(* Logix 5000 project; controller POA Emulate 5570 rev 30.12; software revision 30.00; part 6 of 6 *)
(* tags used below, declared in another part *)
   UOWHF_Add_c : DINT;
   UOWHF_i : DINT;
   UOWHF_InputLen : DINT;
   UOWHF_InputMaxInd : DINT;
   UOWHF_Msg : DINT[17];
   UOWHF_OutputMaxInd : DINT;
   UOWHF_Result : DINT[17];
   UOWHF_Vary_BlkNum : DINT;
   UOWHF_Vary_i : DINT;
   UOWHF_Vary_j : DINT;
   UOWHF_Vary_Message : DINT[3000];
   UOWHF_Vary_MsgLen : DINT;
   UOWHF_Vary_z : DINT;
   UOWHF_VaryLen : DINT;
   UOWHF_Ver : DINT;
(* MainProgram, continued *)

   		UOWHF_Result[0].31:=0;
   		UOWHF_Result[1]:=UOWHF_Result[1] + 1000119182+UOWHF_Add_c;
   		UOWHF_Add_c.1:=UOWHF_Result[1].31;
   		UOWHF_Result[1].31:=0;
   		UOWHF_Result[2]:=UOWHF_Result[2] + 1408193498+UOWHF_Add_c;
   		UOWHF_Add_c.2:=UOWHF_Result[2].31;
   		UOWHF_Result[2].31:=0;
   		UOWHF_Result[3]:=UOWHF_Result[3] + 758141530+UOWHF_Add_c;
   		UOWHF_Add_c.3:=UOWHF_Result[3].31;
   		UOWHF_Result[3].31:=0;
   		UOWHF_Result[4]:=UOWHF_Result[4] + 113758068+UOWHF_Add_c;
   		UOWHF_Add_c.4:=UOWHF_Result[4].31;
   		UOWHF_Result[4].31:=0;
   	End_If;
   	If UOWHF_Msg[7].[27] Then
   		UOWHF_Result[0]:=UOWHF_Result[0] + 86421407+UOWHF_Add_c;
   		UOWHF_Add_c.0:=UOWHF_Result[0].31;
   		UOWHF_Result[0].31:=0;
   		UOWHF_Result[1]:=UOWHF_Result[1] + 209732804+UOWHF_Add_c;
   		UOWHF_Add_c.1:=UOWHF_Result[1].31;
   		UOWHF_Result[1].31:=0;
   		UOWHF_Result[2]:=UOWHF_Result[2] + 502288861+UOWHF_Add_c;
   		UOWHF_Add_c.2:=UOWHF_Result[2].31;
   		UOWHF_Result[2].31:=0;
   		UOWHF_Result[3]:=UOWHF_Result[3] + 1399545115+UOWHF_Add_c;
   		UOWHF_Add_c.3:=UOWHF_Result[3].31;
   		UOWHF_Result[3].31:=0;
   		UOWHF_Result[4]:=UOWHF_Result[4] + 871725095+UOWHF_Add_c;
   		UOWHF_Add_c.4:=UOWHF_Result[4].31;
   		UOWHF_Result[4].31:=0;
   	End_If;
   	If UOWHF_Msg[7].[28] Then
   		UOWHF_Result[0]:=UOWHF_Result[0] + 2145748906+UOWHF_Add_c;
   		UOWHF_Add_c.0:=UOWHF_Result[0].31;
   		UOWHF_Result[0].31:=0;
   		UOWHF_Result[1]:=UOWHF_Result[1] + 750367767+UOWHF_Add_c;
   		UOWHF_Add_c.1:=UOWHF_Result[1].31;
   		UOWHF_Result[1].31:=0;
   		UOWHF_Result[2]:=UOWHF_Result[2] + 52958798+UOWHF_Add_c;
   		UOWHF_Add_c.2:=UOWHF_Result[2].31;
   		UOWHF_Result[2].31:=0;
   		UOWHF_Result[3]:=UOWHF_Result[3] + 299422686+UOWHF_Add_c;
   		UOWHF_Add_c.3:=UOWHF_Result[3].31;
   		UOWHF_Result[3].31:=0;
   		UOWHF_Result[4]:=UOWHF_Result[4] + 308572882+UOWHF_Add_c;
   		UOWHF_Add_c.4:=UOWHF_Result[4].31;
   		UOWHF_Result[4].31:=0;
   	End_If;
   	If UOWHF_Msg[7].[29] Then
   		UOWHF_Result[0]:=UOWHF_Result[0] + 470166861+UOWHF_Add_c;
   		UOWHF_Add_c.0:=UOWHF_Result[0].31;
   		UOWHF_Result[0].31:=0;
   		UOWHF_Result[1]:=UOWHF_Result[1] + 415982775+UOWHF_Add_c;
   		UOWHF_Add_c.1:=UOWHF_Result[1].31;
   		UOWHF_Result[1].31:=0;
   		UOWHF_Result[2]:=UOWHF_Result[2] + 1958329993+UOWHF_Add_c;
   		UOWHF_Add_c.2:=UOWHF_Result[2].31;
   		UOWHF_Result[2].31:=0;
   		UOWHF_Result[3]:=UOWHF_Result[3] + 1087899847+UOWHF_Add_c;
   		UOWHF_Add_c.3:=UOWHF_Result[3].31;
   		UOWHF_Result[3].31:=0;
   		UOWHF_Result[4]:=UOWHF_Result[4] + 290620487+UOWHF_Add_c;
   		UOWHF_Add_c.4:=UOWHF_Result[4].31;
   		UOWHF_Result[4].31:=0;
   	End_If;
   	If UOWHF_Msg[7].[30] Then
   		UOWHF_Result[0]:=UOWHF_Result[0] + 1272966154+UOWHF_Add_c;
   		UOWHF_Add_c.0:=UOWHF_Result[0].31;
   		UOWHF_Result[0].31:=0;
   		UOWHF_Result[1]:=UOWHF_Result[1] + 1453902280+UOWHF_Add_c;
   		UOWHF_Add_c.1:=UOWHF_Result[1].31;
   		UOWHF_Result[1].31:=0;
   		UOWHF_Result[2]:=UOWHF_Result[2] + 39192907+UOWHF_Add_c;
   		UOWHF_Add_c.2:=UOWHF_Result[2].31;
   		UOWHF_Result[2].31:=0;
   		UOWHF_Result[3]:=UOWHF_Result[3] + 1885566212+UOWHF_Add_c;
   		UOWHF_Add_c.3:=UOWHF_Result[3].31;
   		UOWHF_Result[3].31:=0;
   		UOWHF_Result[4]:=UOWHF_Result[4] + 542596261+UOWHF_Add_c;
   		UOWHF_Add_c.4:=UOWHF_Result[4].31;
   		UOWHF_Result[4].31:=0;
   	End_If;
   	If UOWHF_Msg[7].[31] Then
   		UOWHF_Result[0]:=UOWHF_Result[0] + 1141795178+UOWHF_Add_c;
   		UOWHF_Add_c.0:=UOWHF_Result[0].31;
   		UOWHF_Result[0].31:=0;
   		UOWHF_Result[1]:=UOWHF_Result[1] + 2035392703+UOWHF_Add_c;
   		UOWHF_Add_c.1:=UOWHF_Result[1].31;
   		UOWHF_Result[1].31:=0;
   		UOWHF_Result[2]:=UOWHF_Result[2] + 1548772702+UOWHF_Add_c;
   		UOWHF_Add_c.2:=UOWHF_Result[2].31;
   		UOWHF_Result[2].31:=0;
   		UOWHF_Result[3]:=UOWHF_Result[3] + 1915397606+UOWHF_Add_c;
   		UOWHF_Add_c.3:=UOWHF_Result[3].31;
   		UOWHF_Result[3].31:=0;
   		UOWHF_Result[4]:=UOWHF_Result[4] + 1247475076+UOWHF_Add_c;
   		UOWHF_Add_c.4:=UOWHF_Result[4].31;
   		UOWHF_Result[4].31:=0;
   	End_If;
   	UOWHF_Result[UOWHF_OutputMaxInd]:=UOWHF_Result[UOWHF_OutputMaxInd] and 16#F; //clear high bit
END_ROUTINE

ROUTINE UOWHF_Init   (* structured text *)
   Case UOWHF_Ver OF
   0:
   	UOWHF_InputLen:=255;  //bits of input.
   	UOWHF_InputMaxInd:=8;  //maximum index for dints which store the bits of input.
    	For UOWHF_i:=0 to UOWHF_InputMaxInd by 1 do
   		UOWHF_Result[UOWHF_i]:=0;
   	End_For;
   1:
   	UOWHF_InputLen:= 383;
   	UOWHF_InputMaxInd:=12;  //maximum index for array.
    	For UOWHF_i:=0 to UOWHF_InputMaxInd by 1 do
   		UOWHF_Result[UOWHF_i]:=0;
   	End_For;
   2:
   	UOWHF_InputLen:= 511;
   	UOWHF_InputMaxInd:=16;  //maximum index for array.
   	 For UOWHF_i:=0 to UOWHF_InputMaxInd by 1 do
   		UOWHF_Result[UOWHF_i]:=0;
   	End_For;
   End_Case;
   
   UOWHF_OutputMaxInd := UOWHF_InputMaxInd/2;
END_ROUTINE

ROUTINE UOWHF_Vary   (* structured text *)
   
   
   JSR(UOWHF_Init);
   
   
   
   UOWHF_VaryLen:=(UOWHF_Vary_MsgLen+1) MOD (UOWHF_OutputMaxInd+1);
   If UOWHF_VaryLen<>0 Then
   	UOWHF_VaryLen:=UOWHF_OutputMaxInd+1 - UOWHF_VaryLen;
   
   	//pad 1 if neccessary
   	For UOWHF_Vary_i:=UOWHF_Vary_MsgLen+1 to UOWHF_Vary_MsgLen+UOWHF_VaryLen by 1 Do
   
   		UOWHF_Vary_Message[UOWHF_Vary_i]:=65535;
   
   	End_For;
   	UOWHF_Vary_MsgLen:=UOWHF_Vary_MsgLen+UOWHF_VaryLen;
   End_if;
   
   
   UOWHF_Vary_BlkNum:= (UOWHF_Vary_MsgLen+1)/(UOWHF_OutputMaxInd+1)-1 ;
   
   For UOWHF_Vary_i:=0 to UOWHF_InputMaxInd by 1 Do
   	UOWHF_Msg[UOWHF_Vary_i]:=UOWHF_Vary_Message[UOWHF_Vary_i];
   End_For;
   JSR(UOWHF);
   
   UOWHF_Vary_z:=UOWHF_InputMaxInd+1;
   For UOWHF_Vary_i:=2 to UOWHF_Vary_BlkNum by 1 Do
   
   	For UOWHF_Vary_j:=0 to UOWHF_OutputMaxInd by 1 Do
   		UOWHF_Msg[UOWHF_Vary_j]:=UOWHF_Vary_Message[UOWHF_Vary_z+UOWHF_Vary_j];
   		UOWHF_Msg[UOWHF_Vary_j+UOWHF_OutputMaxInd+1]:=UOWHF_Result[UOWHF_Vary_j];
   	End_For;
   	JSR(UOWHF);
   	UOWHF_Vary_z:=UOWHF_Vary_z+UOWHF_OutputMaxInd+1;
   End_For;
   
   
   
END_ROUTINE
END_PROGRAM
